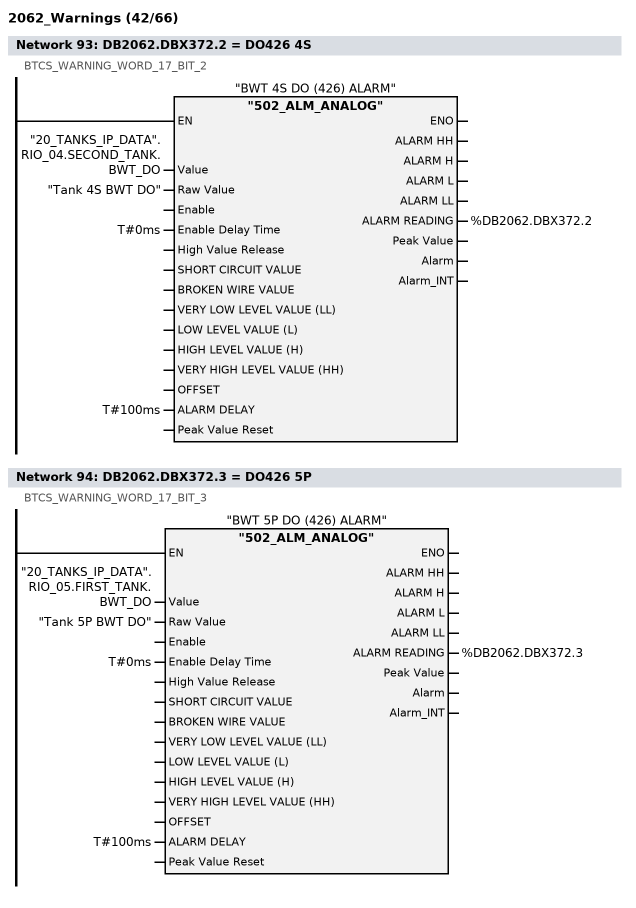
   RUNG wire#powerrail
      "BWT 4S DO (426) ALARM"(Value := "20_TANKS_IP_DATA".RIO_04.SECOND_TANK.BWT_DO, "Raw Value" := "Tank 4S BWT DO", Enable :=, "Enable Delay Time" := T#0ms, "High Value Release" :=, "SHORT CIRCUIT VALUE" :=, "BROKEN WIRE VALUE" :=, "VERY LOW LEVEL VALUE (LL)" :=, "LOW LEVEL VALUE (L)" :=, "HIGH LEVEL VALUE (H)" :=, "VERY HIGH LEVEL VALUE (HH)" :=, OFFSET :=, "ALARM DELAY" := T#100ms, "Peak Value Reset" :=, "ALARM HH" =>, "ALARM H" =>, "ALARM L" =>, "ALARM LL" =>, "ALARM READING" => %DB2062.DBX372.2, "Peak Value" =>, Alarm =>, Alarm_INT =>)
   END_RUNG
   // the same network as SCL:
   "BWT 4S DO (426) ALARM"(Value := "20_TANKS_IP_DATA".RIO_04.SECOND_TANK.BWT_DO,   // "502_ALM_ANALOG"
                           "Raw Value" := "Tank 4S BWT DO",
                           "Enable Delay Time" := T#0ms,
                           "ALARM DELAY" := T#100ms,
                           "ALARM READING" => %DB2062.DBX372.2);
END_REGION

REGION Network 94: DB2062.DBX372.3 = DO426 5P
   // BTCS_WARNING_WORD_17_BIT_3
   RUNG wire#powerrail
      "BWT 5P DO (426) ALARM"(Value := "20_TANKS_IP_DATA".RIO_05.FIRST_TANK.BWT_DO, "Raw Value" := "Tank 5P BWT DO", Enable :=, "Enable Delay Time" := T#0ms, "High Value Release" :=, "SHORT CIRCUIT VALUE" :=, "BROKEN WIRE VALUE" :=, "VERY LOW LEVEL VALUE (LL)" :=, "LOW LEVEL VALUE (L)" :=, "HIGH LEVEL VALUE (H)" :=, "VERY HIGH LEVEL VALUE (HH)" :=, OFFSET :=, "ALARM DELAY" := T#100ms, "Peak Value Reset" :=, "ALARM HH" =>, "ALARM H" =>, "ALARM L" =>, "ALARM LL" =>, "ALARM READING" => %DB2062.DBX372.3, "Peak Value" =>, Alarm =>, Alarm_INT =>)
   END_RUNG
   // the same network as SCL:
   "BWT 5P DO (426) ALARM"(Value := "20_TANKS_IP_DATA".RIO_05.FIRST_TANK.BWT_DO,   // "502_ALM_ANALOG"
                           "Raw Value" := "Tank 5P BWT DO",
                           "Enable Delay Time" := T#0ms,
                           "ALARM DELAY" := T#100ms,
                           "ALARM READING" => %DB2062.DBX372.3);
END_REGION

REGION Network 95: DB2062.DBX372.4 = DO426 5S
   // BTCS_WARNING_WORD_17_BIT_4
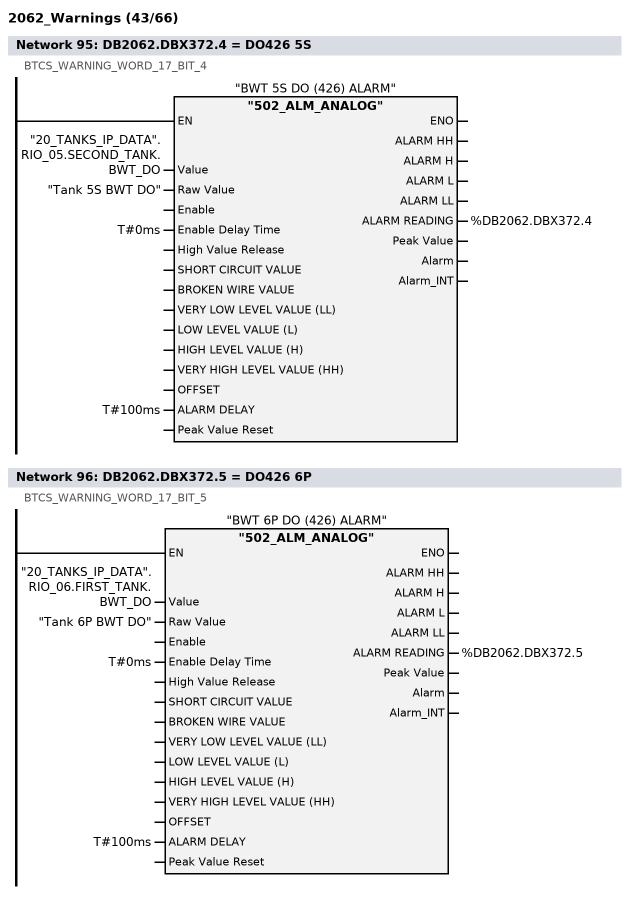
   RUNG wire#powerrail
      "BWT 5S DO (426) ALARM"(Value := "20_TANKS_IP_DATA".RIO_05.SECOND_TANK.BWT_DO, "Raw Value" := "Tank 5S BWT DO", Enable :=, "Enable Delay Time" := T#0ms, "High Value Release" :=, "SHORT CIRCUIT VALUE" :=, "BROKEN WIRE VALUE" :=, "VERY LOW LEVEL VALUE (LL)" :=, "LOW LEVEL VALUE (L)" :=, "HIGH LEVEL VALUE (H)" :=, "VERY HIGH LEVEL VALUE (HH)" :=, OFFSET :=, "ALARM DELAY" := T#100ms, "Peak Value Reset" :=, "ALARM HH" =>, "ALARM H" =>, "ALARM L" =>, "ALARM LL" =>, "ALARM READING" => %DB2062.DBX372.4, "Peak Value" =>, Alarm =>, Alarm_INT =>)
   END_RUNG
   // the same network as SCL:
   "BWT 5S DO (426) ALARM"(Value := "20_TANKS_IP_DATA".RIO_05.SECOND_TANK.BWT_DO,   // "502_ALM_ANALOG"
                           "Raw Value" := "Tank 5S BWT DO",
                           "Enable Delay Time" := T#0ms,
                           "ALARM DELAY" := T#100ms,
                           "ALARM READING" => %DB2062.DBX372.4);
END_REGION

REGION Network 96: DB2062.DBX372.5 = DO426 6P
   // BTCS_WARNING_WORD_17_BIT_5
   RUNG wire#powerrail
      "BWT 6P DO (426) ALARM"(Value := "20_TANKS_IP_DATA".RIO_06.FIRST_TANK.BWT_DO, "Raw Value" := "Tank 6P BWT DO", Enable :=, "Enable Delay Time" := T#0ms, "High Value Release" :=, "SHORT CIRCUIT VALUE" :=, "BROKEN WIRE VALUE" :=, "VERY LOW LEVEL VALUE (LL)" :=, "LOW LEVEL VALUE (L)" :=, "HIGH LEVEL VALUE (H)" :=, "VERY HIGH LEVEL VALUE (HH)" :=, OFFSET :=, "ALARM DELAY" := T#100ms, "Peak Value Reset" :=, "ALARM HH" =>, "ALARM H" =>, "ALARM L" =>, "ALARM LL" =>, "ALARM READING" => %DB2062.DBX372.5, "Peak Value" =>, Alarm =>, Alarm_INT =>)
   END_RUNG
   // the same network as SCL:
   "BWT 6P DO (426) ALARM"(Value := "20_TANKS_IP_DATA".RIO_06.FIRST_TANK.BWT_DO,   // "502_ALM_ANALOG"
                           "Raw Value" := "Tank 6P BWT DO",
                           "Enable Delay Time" := T#0ms,
                           "ALARM DELAY" := T#100ms,
                           "ALARM READING" => %DB2062.DBX372.5);
END_REGION

REGION Network 97: DB2062.DBX372.6 = DO426 6S
   // BTCS_WARNING_WORD_17_BIT_6
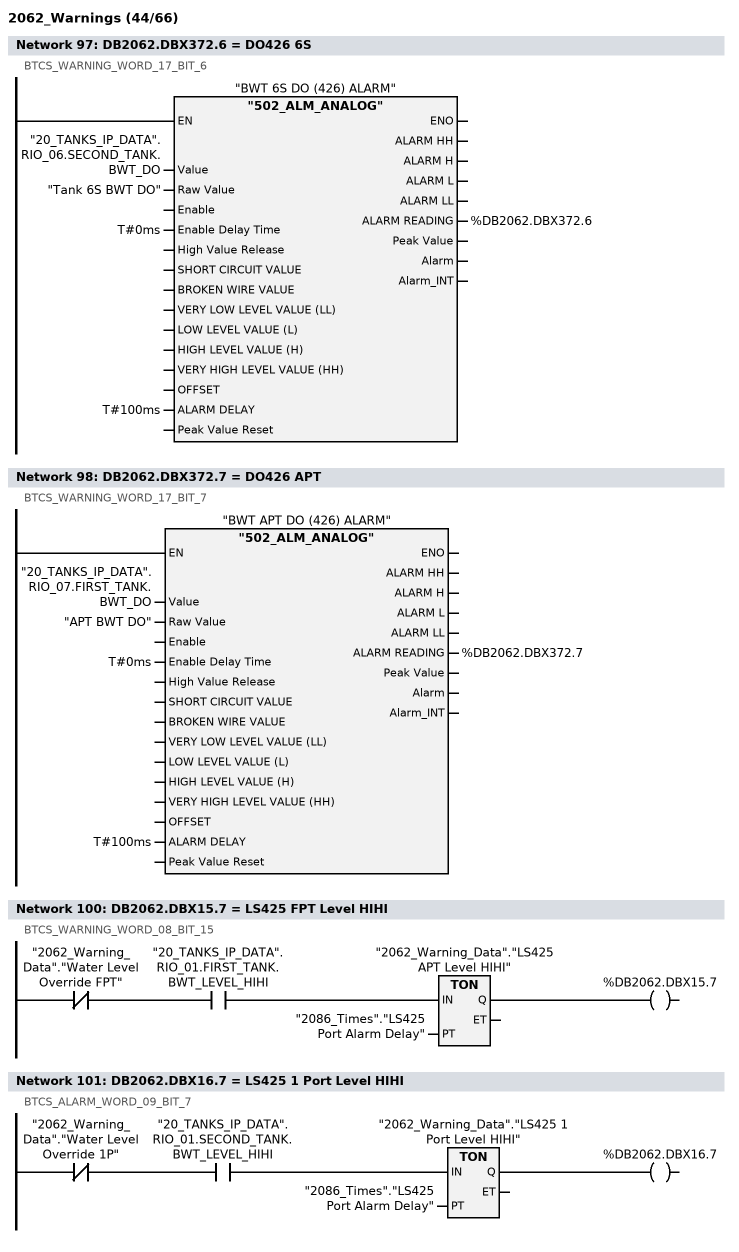
   RUNG wire#powerrail
      "BWT 6S DO (426) ALARM"(Value := "20_TANKS_IP_DATA".RIO_06.SECOND_TANK.BWT_DO, "Raw Value" := "Tank 6S BWT DO", Enable :=, "Enable Delay Time" := T#0ms, "High Value Release" :=, "SHORT CIRCUIT VALUE" :=, "BROKEN WIRE VALUE" :=, "VERY LOW LEVEL VALUE (LL)" :=, "LOW LEVEL VALUE (L)" :=, "HIGH LEVEL VALUE (H)" :=, "VERY HIGH LEVEL VALUE (HH)" :=, OFFSET :=, "ALARM DELAY" := T#100ms, "Peak Value Reset" :=, "ALARM HH" =>, "ALARM H" =>, "ALARM L" =>, "ALARM LL" =>, "ALARM READING" => %DB2062.DBX372.6, "Peak Value" =>, Alarm =>, Alarm_INT =>)
   END_RUNG
   // the same network as SCL:
   "BWT 6S DO (426) ALARM"(Value := "20_TANKS_IP_DATA".RIO_06.SECOND_TANK.BWT_DO,   // "502_ALM_ANALOG"
                           "Raw Value" := "Tank 6S BWT DO",
                           "Enable Delay Time" := T#0ms,
                           "ALARM DELAY" := T#100ms,
                           "ALARM READING" => %DB2062.DBX372.6);
END_REGION

REGION Network 98: DB2062.DBX372.7 = DO426 APT
   // BTCS_WARNING_WORD_17_BIT_7
   RUNG wire#powerrail
      "BWT APT DO (426) ALARM"(Value := "20_TANKS_IP_DATA".RIO_07.FIRST_TANK.BWT_DO, "Raw Value" := "APT BWT DO", Enable :=, "Enable Delay Time" := T#0ms, "High Value Release" :=, "SHORT CIRCUIT VALUE" :=, "BROKEN WIRE VALUE" :=, "VERY LOW LEVEL VALUE (LL)" :=, "LOW LEVEL VALUE (L)" :=, "HIGH LEVEL VALUE (H)" :=, "VERY HIGH LEVEL VALUE (HH)" :=, OFFSET :=, "ALARM DELAY" := T#100ms, "Peak Value Reset" :=, "ALARM HH" =>, "ALARM H" =>, "ALARM L" =>, "ALARM LL" =>, "ALARM READING" => %DB2062.DBX372.7, "Peak Value" =>, Alarm =>, Alarm_INT =>)
   END_RUNG
   // the same network as SCL:
   "BWT APT DO (426) ALARM"(Value := "20_TANKS_IP_DATA".RIO_07.FIRST_TANK.BWT_DO,   // "502_ALM_ANALOG"
                           "Raw Value" := "APT BWT DO",
                           "Enable Delay Time" := T#0ms,
                           "ALARM DELAY" := T#100ms,
                           "ALARM READING" => %DB2062.DBX372.7);
END_REGION

REGION Network 100: DB2062.DBX15.7 = LS425 FPT Level HIHI
   // BTCS_WARNING_WORD_08_BIT_15
   "2062_Warning_Data"."LS425 APT Level HIHI".TON(IN := NOT "2062_Warning_Data"."Water Level Override FPT" AND "20_TANKS_IP_DATA".RIO_01.FIRST_TANK.BWT_LEVEL_HIHI,
                           PT := "2086_Times"."LS425 Port Alarm Delay");
   %DB2062.DBX15.7 := "2062_Warning_Data"."LS425 APT Level HIHI".Q;
END_REGION

REGION Network 101: DB2062.DBX16.7 = LS425 1 Port Level HIHI
   // BTCS_ALARM_WORD_09_BIT_7
   "2062_Warning_Data"."LS425 1 Port Level HIHI".TON(IN := NOT "2062_Warning_Data"."Water Level Override 1P" AND "20_TANKS_IP_DATA".RIO_01.SECOND_TANK.BWT_LEVEL_HIHI,
                           PT := "2086_Times"."LS425 Port Alarm Delay");
   %DB2062.DBX16.7 := "2062_Warning_Data"."LS425 1 Port Level HIHI".Q;
END_REGION

REGION Network 102: DB2062.DBX14.2 = LS425 1 Starboard Level HIHI
   // BTCS_ALARM_WORD_08_BIT_2
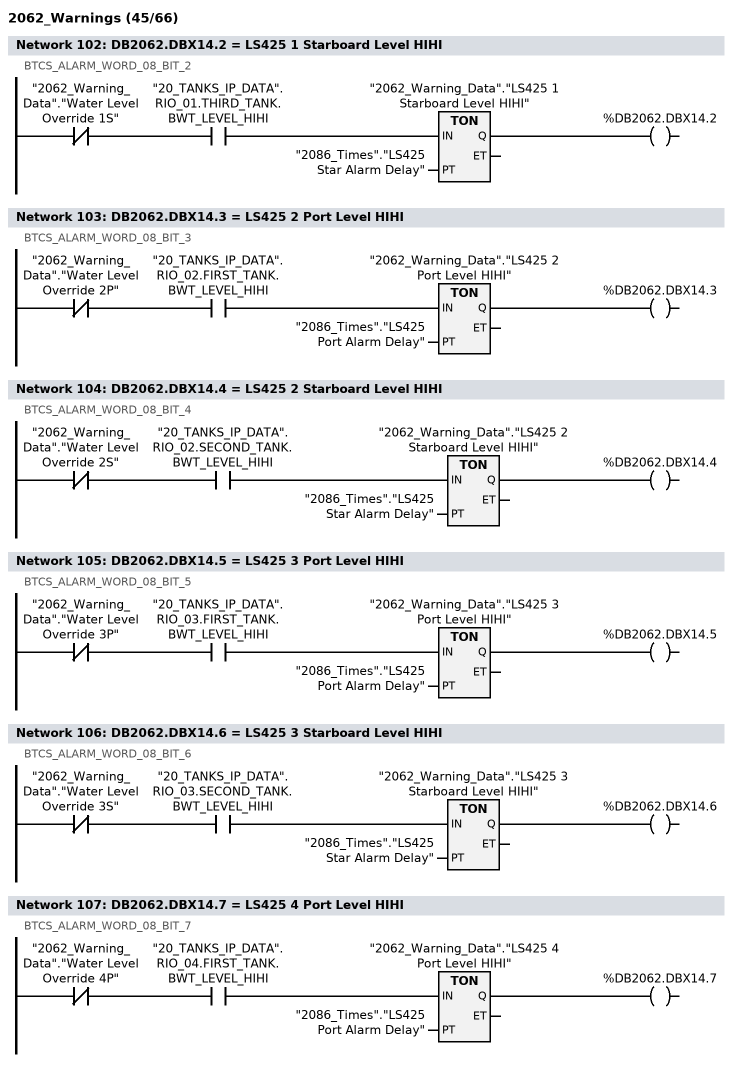
   "2062_Warning_Data"."LS425 1 Starboard Level HIHI".TON(IN := NOT "2062_Warning_Data"."Water Level Override 1S" AND "20_TANKS_IP_DATA".RIO_01.THIRD_TANK.BWT_LEVEL_HIHI,
                           PT := "2086_Times"."LS425 Star Alarm Delay");
   %DB2062.DBX14.2 := "2062_Warning_Data"."LS425 1 Starboard Level HIHI".Q;
END_REGION

REGION Network 103: DB2062.DBX14.3 = LS425 2 Port Level HIHI
   // BTCS_ALARM_WORD_08_BIT_3
   "2062_Warning_Data"."LS425 2 Port Level HIHI".TON(IN := NOT "2062_Warning_Data"."Water Level Override 2P" AND "20_TANKS_IP_DATA".RIO_02.FIRST_TANK.BWT_LEVEL_HIHI,
                           PT := "2086_Times"."LS425 Port Alarm Delay");
   %DB2062.DBX14.3 := "2062_Warning_Data"."LS425 2 Port Level HIHI".Q;
END_REGION

REGION Network 104: DB2062.DBX14.4 = LS425 2 Starboard Level HIHI
   // BTCS_ALARM_WORD_08_BIT_4
   "2062_Warning_Data"."LS425 2 Starboard Level HIHI".TON(IN := NOT "2062_Warning_Data"."Water Level Override 2S" AND "20_TANKS_IP_DATA".RIO_02.SECOND_TANK.BWT_LEVEL_HIHI,
                           PT := "2086_Times"."LS425 Star Alarm Delay");
   %DB2062.DBX14.4 := "2062_Warning_Data"."LS425 2 Starboard Level HIHI".Q;
END_REGION

REGION Network 105: DB2062.DBX14.5 = LS425 3 Port Level HIHI
   // BTCS_ALARM_WORD_08_BIT_5
   "2062_Warning_Data"."LS425 3 Port Level HIHI".TON(IN := NOT "2062_Warning_Data"."Water Level Override 3P" AND "20_TANKS_IP_DATA".RIO_03.FIRST_TANK.BWT_LEVEL_HIHI,
                           PT := "2086_Times"."LS425 Port Alarm Delay");
   %DB2062.DBX14.5 := "2062_Warning_Data"."LS425 3 Port Level HIHI".Q;
END_REGION

REGION Network 106: DB2062.DBX14.6 = LS425 3 Starboard Level HIHI
   // BTCS_ALARM_WORD_08_BIT_6
   "2062_Warning_Data"."LS425 3 Starboard Level HIHI".TON(IN := NOT "2062_Warning_Data"."Water Level Override 3S" AND "20_TANKS_IP_DATA".RIO_03.SECOND_TANK.BWT_LEVEL_HIHI,
                           PT := "2086_Times"."LS425 Star Alarm Delay");
   %DB2062.DBX14.6 := "2062_Warning_Data"."LS425 3 Starboard Level HIHI".Q;
END_REGION

REGION Network 107: DB2062.DBX14.7 = LS425 4 Port Level HIHI
   // BTCS_ALARM_WORD_08_BIT_7
   "2062_Warning_Data"."LS425 4 Port Level HIHI".TON(IN := NOT "2062_Warning_Data"."Water Level Override 4P" AND "20_TANKS_IP_DATA".RIO_04.FIRST_TANK.BWT_LEVEL_HIHI,
                           PT := "2086_Times"."LS425 Port Alarm Delay");
   %DB2062.DBX14.7 := "2062_Warning_Data"."LS425 4 Port Level HIHI".Q;
END_REGION

REGION Network 108: DB2062.DBX15.0 = LS425 4 Starboard Level HIHI
   // BTCS_ALARM_WORD_08_BIT_8
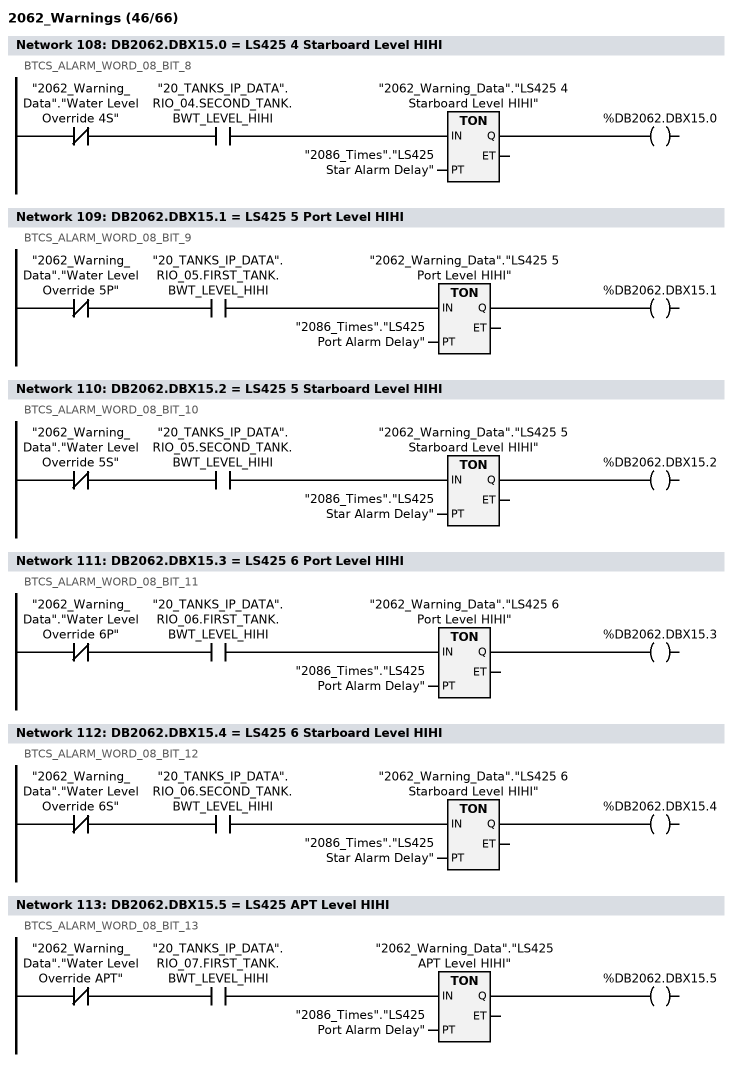
   "2062_Warning_Data"."LS425 4 Starboard Level HIHI".TON(IN := NOT "2062_Warning_Data"."Water Level Override 4S" AND "20_TANKS_IP_DATA".RIO_04.SECOND_TANK.BWT_LEVEL_HIHI,
                           PT := "2086_Times"."LS425 Star Alarm Delay");
   %DB2062.DBX15.0 := "2062_Warning_Data"."LS425 4 Starboard Level HIHI".Q;
END_REGION

REGION Network 109: DB2062.DBX15.1 = LS425 5 Port Level HIHI
   // BTCS_ALARM_WORD_08_BIT_9
   "2062_Warning_Data"."LS425 5 Port Level HIHI".TON(IN := NOT "2062_Warning_Data"."Water Level Override 5P" AND "20_TANKS_IP_DATA".RIO_05.FIRST_TANK.BWT_LEVEL_HIHI,
                           PT := "2086_Times"."LS425 Port Alarm Delay");
   %DB2062.DBX15.1 := "2062_Warning_Data"."LS425 5 Port Level HIHI".Q;
END_REGION

REGION Network 110: DB2062.DBX15.2 = LS425 5 Starboard Level HIHI
   // BTCS_ALARM_WORD_08_BIT_10
   "2062_Warning_Data"."LS425 5 Starboard Level HIHI".TON(IN := NOT "2062_Warning_Data"."Water Level Override 5S" AND "20_TANKS_IP_DATA".RIO_05.SECOND_TANK.BWT_LEVEL_HIHI,
                           PT := "2086_Times"."LS425 Star Alarm Delay");
   %DB2062.DBX15.2 := "2062_Warning_Data"."LS425 5 Starboard Level HIHI".Q;
END_REGION

REGION Network 111: DB2062.DBX15.3 = LS425 6 Port Level HIHI
   // BTCS_ALARM_WORD_08_BIT_11
   "2062_Warning_Data"."LS425 6 Port Level HIHI".TON(IN := NOT "2062_Warning_Data"."Water Level Override 6P" AND "20_TANKS_IP_DATA".RIO_06.FIRST_TANK.BWT_LEVEL_HIHI,
                           PT := "2086_Times"."LS425 Port Alarm Delay");
   %DB2062.DBX15.3 := "2062_Warning_Data"."LS425 6 Port Level HIHI".Q;
END_REGION

REGION Network 112: DB2062.DBX15.4 = LS425 6 Starboard Level HIHI
   // BTCS_ALARM_WORD_08_BIT_12
   "2062_Warning_Data"."LS425 6 Starboard Level HIHI".TON(IN := NOT "2062_Warning_Data"."Water Level Override 6S" AND "20_TANKS_IP_DATA".RIO_06.SECOND_TANK.BWT_LEVEL_HIHI,
                           PT := "2086_Times"."LS425 Star Alarm Delay");
   %DB2062.DBX15.4 := "2062_Warning_Data"."LS425 6 Starboard Level HIHI".Q;
END_REGION

REGION Network 113: DB2062.DBX15.5 = LS425 APT Level HIHI
   // BTCS_ALARM_WORD_08_BIT_13
   "2062_Warning_Data"."LS425 APT Level HIHI".TON(IN := NOT "2062_Warning_Data"."Water Level Override APT" AND "20_TANKS_IP_DATA".RIO_07.FIRST_TANK.BWT_LEVEL_HIHI,
                           PT := "2086_Times"."LS425 Port Alarm Delay");
   %DB2062.DBX15.5 := "2062_Warning_Data"."LS425 APT Level HIHI".Q;
END_REGION

REGION Network 115: DB2062.DBX16.0 = PS436 RIO1 Tank Group Pressure HIHI
   // BTCS_ALARM_WORD_09_BIT_0
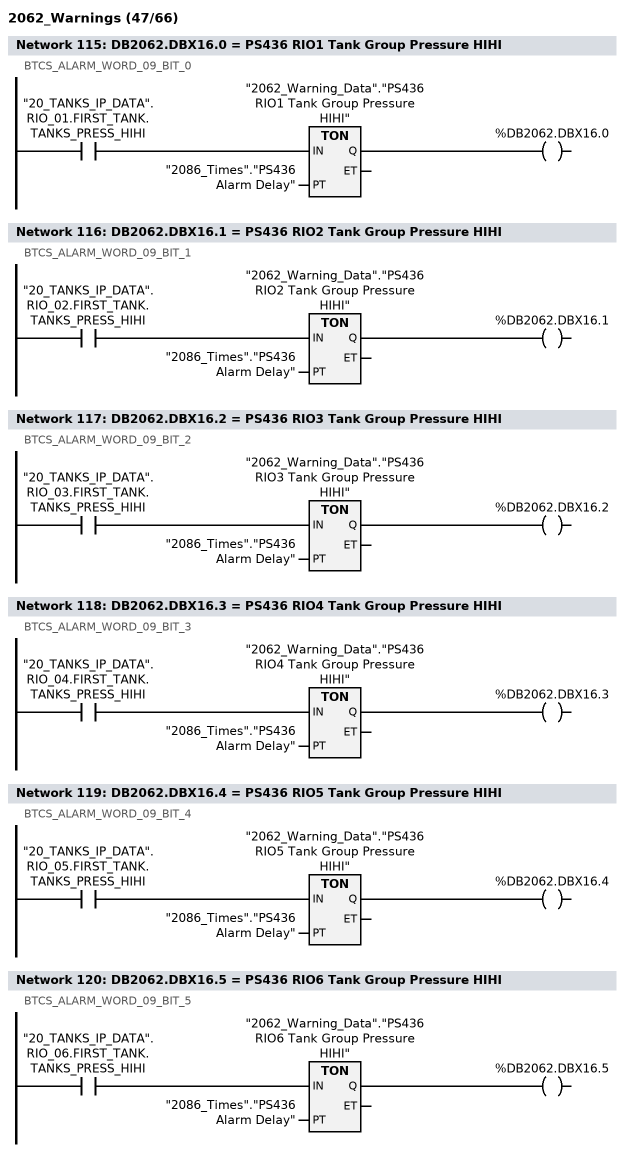
   "2062_Warning_Data"."PS436 RIO1 Tank Group Pressure HIHI".TON(IN := "20_TANKS_IP_DATA".RIO_01.FIRST_TANK.TANKS_PRESS_HIHI,
                           PT := "2086_Times"."PS436 Alarm Delay");
   %DB2062.DBX16.0 := "2062_Warning_Data"."PS436 RIO1 Tank Group Pressure HIHI".Q;
END_REGION

REGION Network 116: DB2062.DBX16.1 = PS436 RIO2 Tank Group Pressure HIHI
   // BTCS_ALARM_WORD_09_BIT_1
   "2062_Warning_Data"."PS436 RIO2 Tank Group Pressure HIHI".TON(IN := "20_TANKS_IP_DATA".RIO_02.FIRST_TANK.TANKS_PRESS_HIHI,
                           PT := "2086_Times"."PS436 Alarm Delay");
   %DB2062.DBX16.1 := "2062_Warning_Data"."PS436 RIO2 Tank Group Pressure HIHI".Q;
END_REGION

REGION Network 117: DB2062.DBX16.2 = PS436 RIO3 Tank Group Pressure HIHI
   // BTCS_ALARM_WORD_09_BIT_2
   "2062_Warning_Data"."PS436 RIO3 Tank Group Pressure HIHI".TON(IN := "20_TANKS_IP_DATA".RIO_03.FIRST_TANK.TANKS_PRESS_HIHI,
                           PT := "2086_Times"."PS436 Alarm Delay");
   %DB2062.DBX16.2 := "2062_Warning_Data"."PS436 RIO3 Tank Group Pressure HIHI".Q;
END_REGION

REGION Network 118: DB2062.DBX16.3 = PS436 RIO4 Tank Group Pressure HIHI
   // BTCS_ALARM_WORD_09_BIT_3
   "2062_Warning_Data"."PS436 RIO4 Tank Group Pressure HIHI".TON(IN := "20_TANKS_IP_DATA".RIO_04.FIRST_TANK.TANKS_PRESS_HIHI,
                           PT := "2086_Times"."PS436 Alarm Delay");
   %DB2062.DBX16.3 := "2062_Warning_Data"."PS436 RIO4 Tank Group Pressure HIHI".Q;
END_REGION

REGION Network 119: DB2062.DBX16.4 = PS436 RIO5 Tank Group Pressure HIHI
   // BTCS_ALARM_WORD_09_BIT_4
   "2062_Warning_Data"."PS436 RIO5 Tank Group Pressure HIHI".TON(IN := "20_TANKS_IP_DATA".RIO_05.FIRST_TANK.TANKS_PRESS_HIHI,
                           PT := "2086_Times"."PS436 Alarm Delay");
   %DB2062.DBX16.4 := "2062_Warning_Data"."PS436 RIO5 Tank Group Pressure HIHI".Q;
END_REGION

REGION Network 120: DB2062.DBX16.5 = PS436 RIO6 Tank Group Pressure HIHI
   // BTCS_ALARM_WORD_09_BIT_5
   "2062_Warning_Data"."PS436 RIO6 Tank Group Pressure HIHI".TON(IN := "20_TANKS_IP_DATA".RIO_06.FIRST_TANK.TANKS_PRESS_HIHI,
                           PT := "2086_Times"."PS436 Alarm Delay");
   %DB2062.DBX16.5 := "2062_Warning_Data"."PS436 RIO6 Tank Group Pressure HIHI".Q;
END_REGION

REGION Network 121: DB2062.DBX16.6 = PS436 RIO7 Tank Group Pressure HIHI
   // BTCS_ALARM_WORD_09_BIT_6
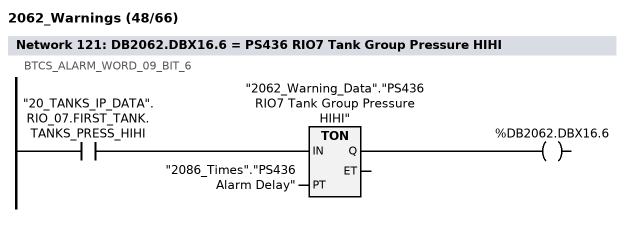
   "2062_Warning_Data"."PS436 RIO7 Tank Group Pressure HIHI".TON(IN := "20_TANKS_IP_DATA".RIO_07.FIRST_TANK.TANKS_PRESS_HIHI,
                           PT := "2086_Times"."PS436 Alarm Delay");
   %DB2062.DBX16.6 := "2062_Warning_Data"."PS436 RIO7 Tank Group Pressure HIHI".Q;
END_REGION

REGION Network 123: Level Override Set
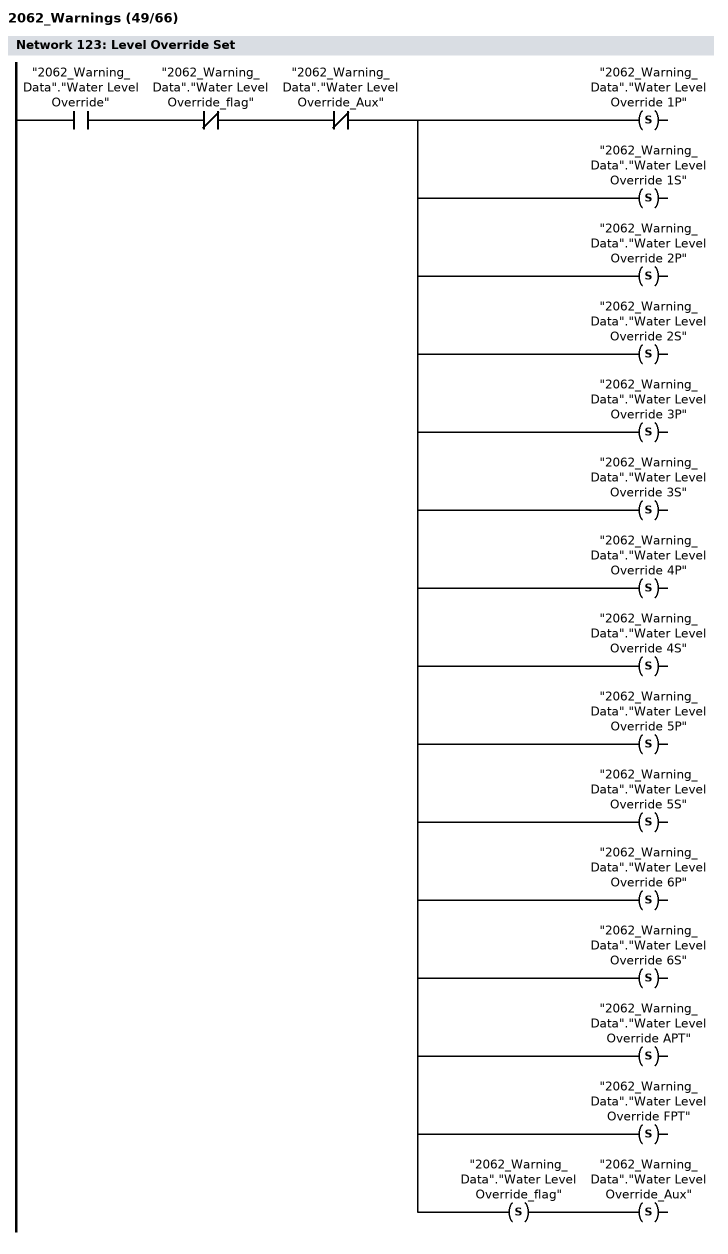
   RUNG wire#powerrail
      Contact( "2062_Warning_Data"."Water Level Override" )
      I_Contact( "2062_Warning_Data"."Water Level Override_flag" )
      I_Contact( "2062_Warning_Data"."Water Level Override_Aux" )
      wire#w1
      S_Coil( "2062_Warning_Data"."Water Level Override 1P" )
   END_RUNG
   RUNG wire#w1
      S_Coil( "2062_Warning_Data"."Water Level Override 1S" )
   END_RUNG
   RUNG wire#w1
      S_Coil( "2062_Warning_Data"."Water Level Override 2P" )
   END_RUNG
   RUNG wire#w1
      S_Coil( "2062_Warning_Data"."Water Level Override 2S" )
   END_RUNG
   RUNG wire#w1
      S_Coil( "2062_Warning_Data"."Water Level Override 3P" )
   END_RUNG
   RUNG wire#w1
      S_Coil( "2062_Warning_Data"."Water Level Override 3S" )
   END_RUNG
   RUNG wire#w1
      S_Coil( "2062_Warning_Data"."Water Level Override 4P" )
   END_RUNG
   RUNG wire#w1
      S_Coil( "2062_Warning_Data"."Water Level Override 4S" )
   END_RUNG
   RUNG wire#w1
      S_Coil( "2062_Warning_Data"."Water Level Override 5P" )
   END_RUNG
   RUNG wire#w1
      S_Coil( "2062_Warning_Data"."Water Level Override 5S" )
   END_RUNG
   RUNG wire#w1
      S_Coil( "2062_Warning_Data"."Water Level Override 6P" )
   END_RUNG
   RUNG wire#w1
      S_Coil( "2062_Warning_Data"."Water Level Override 6S" )
   END_RUNG
   RUNG wire#w1
      S_Coil( "2062_Warning_Data"."Water Level Override APT" )
   END_RUNG
   RUNG wire#w1
      S_Coil( "2062_Warning_Data"."Water Level Override FPT" )
   END_RUNG
   RUNG wire#w1
      S_Coil( "2062_Warning_Data"."Water Level Override_flag" )
      S_Coil( "2062_Warning_Data"."Water Level Override_Aux" )
   END_RUNG
   // the same network as SCL:
   IF "2062_Warning_Data"."Water Level Override" AND NOT "2062_Warning_Data"."Water Level Override_flag" AND NOT "2062_Warning_Data"."Water Level Override_Aux" THEN
       "2062_Warning_Data"."Water Level Override 1P" := TRUE;
       "2062_Warning_Data"."Water Level Override 1S" := TRUE;
       "2062_Warning_Data"."Water Level Override 2P" := TRUE;
       "2062_Warning_Data"."Water Level Override 2S" := TRUE;
       "2062_Warning_Data"."Water Level Override 3P" := TRUE;
       "2062_Warning_Data"."Water Level Override 3S" := TRUE;
       "2062_Warning_Data"."Water Level Override 4P" := TRUE;
       "2062_Warning_Data"."Water Level Override 4S" := TRUE;
       "2062_Warning_Data"."Water Level Override 5P" := TRUE;
       "2062_Warning_Data"."Water Level Override 5S" := TRUE;
       "2062_Warning_Data"."Water Level Override 6P" := TRUE;
       "2062_Warning_Data"."Water Level Override 6S" := TRUE;
       "2062_Warning_Data"."Water Level Override APT" := TRUE;
       "2062_Warning_Data"."Water Level Override FPT" := TRUE;
   END_IF;
   #_w1 := "2062_Warning_Data"."Water Level Override" AND NOT "2062_Warning_Data"."Water Level Override_flag" AND NOT "2062_Warning_Data"."Water Level Override_Aux";
   IF #_w1 THEN
       "2062_Warning_Data"."Water Level Override_flag" := TRUE;
       "2062_Warning_Data"."Water Level Override_Aux" := TRUE;
   END_IF;
END_REGION

REGION Network 124: Level Override Reset
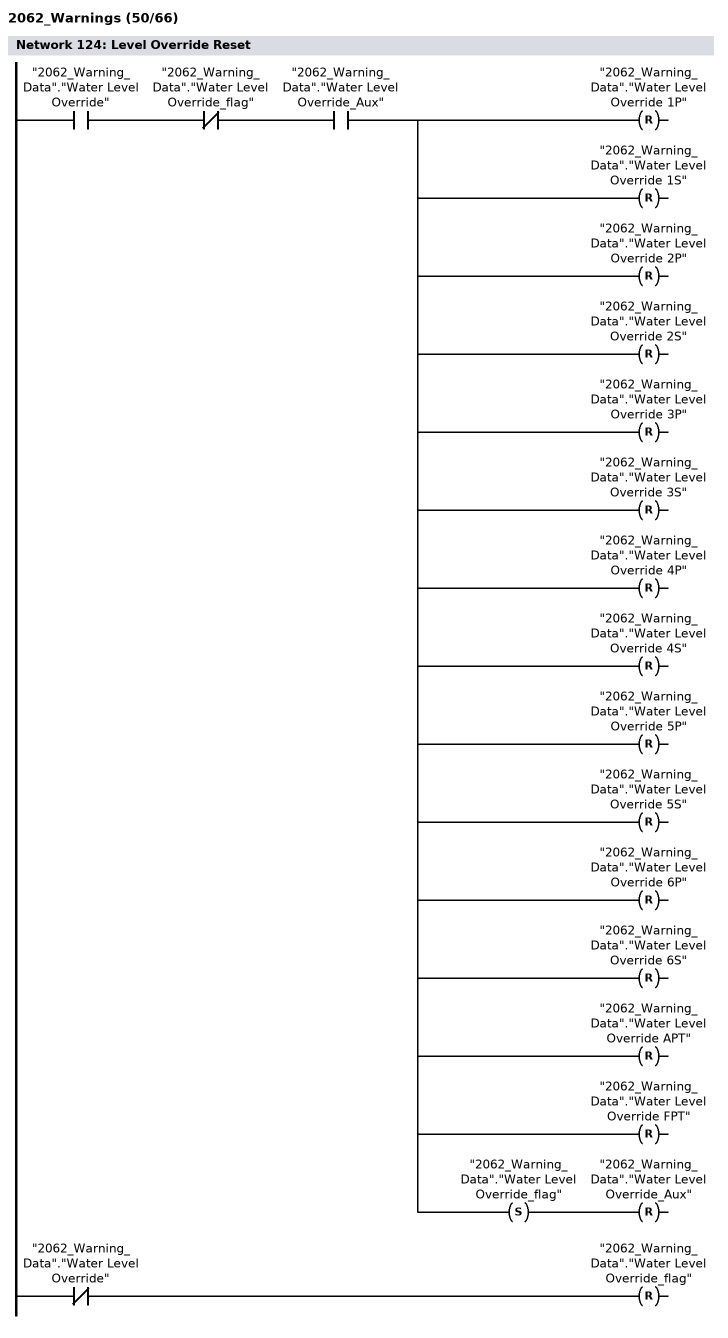
   RUNG wire#powerrail
      Contact( "2062_Warning_Data"."Water Level Override" )
      I_Contact( "2062_Warning_Data"."Water Level Override_flag" )
      Contact( "2062_Warning_Data"."Water Level Override_Aux" )
      wire#w1
      R_Coil( "2062_Warning_Data"."Water Level Override 1P" )
   END_RUNG
   RUNG wire#w1
      R_Coil( "2062_Warning_Data"."Water Level Override 1S" )
   END_RUNG
   RUNG wire#w1
      R_Coil( "2062_Warning_Data"."Water Level Override 2P" )
   END_RUNG
   RUNG wire#w1
      R_Coil( "2062_Warning_Data"."Water Level Override 2S" )
   END_RUNG
   RUNG wire#w1
      R_Coil( "2062_Warning_Data"."Water Level Override 3P" )
   END_RUNG
   RUNG wire#w1
      R_Coil( "2062_Warning_Data"."Water Level Override 3S" )
   END_RUNG
   RUNG wire#w1
      R_Coil( "2062_Warning_Data"."Water Level Override 4P" )
   END_RUNG
   RUNG wire#w1
      R_Coil( "2062_Warning_Data"."Water Level Override 4S" )
   END_RUNG
   RUNG wire#w1
      R_Coil( "2062_Warning_Data"."Water Level Override 5P" )
   END_RUNG
   RUNG wire#w1
      R_Coil( "2062_Warning_Data"."Water Level Override 5S" )
   END_RUNG
   RUNG wire#w1
      R_Coil( "2062_Warning_Data"."Water Level Override 6P" )
   END_RUNG
   RUNG wire#w1
      R_Coil( "2062_Warning_Data"."Water Level Override 6S" )
   END_RUNG
   RUNG wire#w1
      R_Coil( "2062_Warning_Data"."Water Level Override APT" )
   END_RUNG
   RUNG wire#w1
      R_Coil( "2062_Warning_Data"."Water Level Override FPT" )
   END_RUNG
   RUNG wire#w1
      S_Coil( "2062_Warning_Data"."Water Level Override_flag" )
      R_Coil( "2062_Warning_Data"."Water Level Override_Aux" )
   END_RUNG
   RUNG wire#powerrail
      I_Contact( "2062_Warning_Data"."Water Level Override" )
      R_Coil( "2062_Warning_Data"."Water Level Override_flag" )
   END_RUNG
   // the same network as SCL:
   IF "2062_Warning_Data"."Water Level Override" AND NOT "2062_Warning_Data"."Water Level Override_flag" AND "2062_Warning_Data"."Water Level Override_Aux" THEN
       "2062_Warning_Data"."Water Level Override 1P" := FALSE;
       "2062_Warning_Data"."Water Level Override 1S" := FALSE;
       "2062_Warning_Data"."Water Level Override 2P" := FALSE;
       "2062_Warning_Data"."Water Level Override 2S" := FALSE;
       "2062_Warning_Data"."Water Level Override 3P" := FALSE;
       "2062_Warning_Data"."Water Level Override 3S" := FALSE;
       "2062_Warning_Data"."Water Level Override 4P" := FALSE;
       "2062_Warning_Data"."Water Level Override 4S" := FALSE;
       "2062_Warning_Data"."Water Level Override 5P" := FALSE;
       "2062_Warning_Data"."Water Level Override 5S" := FALSE;
       "2062_Warning_Data"."Water Level Override 6P" := FALSE;
       "2062_Warning_Data"."Water Level Override 6S" := FALSE;
       "2062_Warning_Data"."Water Level Override APT" := FALSE;
       "2062_Warning_Data"."Water Level Override FPT" := FALSE;
   END_IF;
   #_w1 := "2062_Warning_Data"."Water Level Override" AND NOT "2062_Warning_Data"."Water Level Override_flag" AND "2062_Warning_Data"."Water Level Override_Aux";
   IF #_w1 THEN
       "2062_Warning_Data"."Water Level Override_flag" := TRUE;
       "2062_Warning_Data"."Water Level Override_Aux" := FALSE;
   END_IF;
   IF NOT "2062_Warning_Data"."Water Level Override" THEN
       "2062_Warning_Data"."Water Level Override_flag" := FALSE;
   END_IF;
END_REGION

REGION Network 125: DB2062.DBX17.0/1 = LT422 FPT Tank Level
   // BTCS_ALARM_WORD_09_BIT_8/9                             14.12
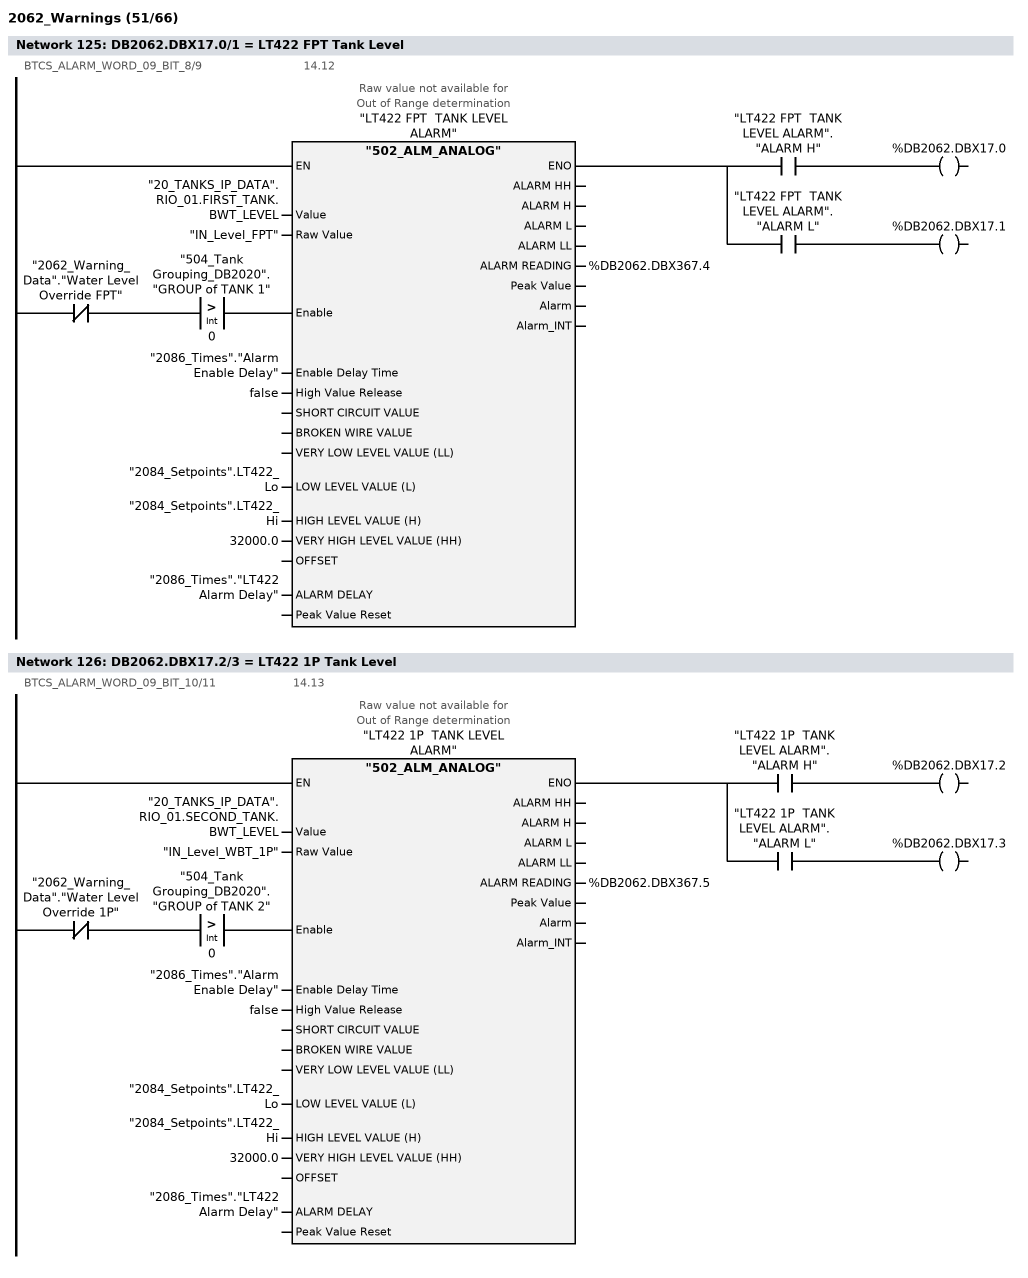
   RUNG wire#powerrail
      "LT422 FPT  TANK LEVEL ALARM"(Enable := wire#w1, Value := "20_TANKS_IP_DATA".RIO_01.FIRST_TANK.BWT_LEVEL, "Raw Value" := "IN_Level_FPT", "Enable Delay Time" := "2086_Times"."Alarm Enable Delay", "High Value Release" := false, "SHORT CIRCUIT VALUE" :=, "BROKEN WIRE VALUE" :=, "VERY LOW LEVEL VALUE (LL)" :=, "LOW LEVEL VALUE (L)" := "2084_Setpoints".LT422_Lo, "HIGH LEVEL VALUE (H)" := "2084_Setpoints".LT422_Hi, "VERY HIGH LEVEL VALUE (HH)" := 32000.0, OFFSET :=, "ALARM DELAY" := "2086_Times"."LT422 Alarm Delay", "Peak Value Reset" :=, "ALARM HH" =>, "ALARM H" =>, "ALARM L" =>, "ALARM LL" =>, "ALARM READING" => %DB2062.DBX367.4, "Peak Value" =>, Alarm =>, Alarm_INT =>)   // Raw value not available for Out of Range determination
      wire#w2
      Contact( "LT422 FPT  TANK LEVEL ALARM"."ALARM H" )
      Coil( %DB2062.DBX17.0 )
   END_RUNG
   RUNG wire#powerrail
      I_Contact( "2062_Warning_Data"."Water Level Override FPT" )
      { S7_Templates := "SrcType := Int" } GT_Contact(in1 := "504_Tank Grouping_DB2020"."GROUP of TANK 1", in2 := 0)
   END_RUNG wire#w1
   RUNG wire#w2
      Contact( "LT422 FPT  TANK LEVEL ALARM"."ALARM L" )
      Coil( %DB2062.DBX17.1 )
   END_RUNG
   // the same network as SCL:
   "LT422 FPT  TANK LEVEL ALARM"(Value := "20_TANKS_IP_DATA".RIO_01.FIRST_TANK.BWT_LEVEL,   // "502_ALM_ANALOG": Raw value not available for Out of Range determination
                           "Raw Value" := "IN_Level_FPT",
                           Enable := NOT "2062_Warning_Data"."Water Level Override FPT" AND ("504_Tank Grouping_DB2020"."GROUP of TANK 1" > 0),
                           "Enable Delay Time" := "2086_Times"."Alarm Enable Delay",
                           "High Value Release" := false,
                           "LOW LEVEL VALUE (L)" := "2084_Setpoints".LT422_Lo,
                           "HIGH LEVEL VALUE (H)" := "2084_Setpoints".LT422_Hi,
                           "VERY HIGH LEVEL VALUE (HH)" := 32000.0,
                           "ALARM DELAY" := "2086_Times"."LT422 Alarm Delay",
                           "ALARM READING" => %DB2062.DBX367.4,
                           ENO => #_w1);
   %DB2062.DBX17.0 := #_w1 AND "LT422 FPT  TANK LEVEL ALARM"."ALARM H";
   %DB2062.DBX17.1 := #_w1 AND "LT422 FPT  TANK LEVEL ALARM"."ALARM L";
END_REGION
